screen "1121_OMACPackTags" 1280x715, template "1xxx_MachineControl"
   TextField "fraStatusPackTags" at 15,15 size 535x225; Text 'Status / Estado:'
   TextField "txtStatusCurUnitMode" at 25,55 size 220x25; Text 'Unit mode current: / Aktuelle Betriebsart: / Modo de unidad actual:'
   TextField "txtStatusCurState" at 25,85 size 220x25; Text 'State current: / Aktueller Zustand: / Corriente del estado'
   TextField "txtStatusCurMachSpeed" at 25,115 size 220x25; Text 'Current machine speed: / Aktuelle Geschwindigkeit'
   TextField "txtStatusCurMachSpeedUnit" at 370,115 size 80x25; Text 'pcs/min / Stck/Min / m/min'
   TextField "txtStatusMachSpeed" at 25,145 size 220x25; Text 'Machine speed: / Maschinengeschwindigkeit: / Velocidad de la máquina:'
   TextField "txtStatusMachSpeedUnit" at 370,145 size 80x25; Text 'pcs/min / Stck/Min / m/min'
   TextField "txtStatusEquipmentInterlockBlocked" at 25,175 size 220x25; Text 'Equip. interlock blocked: / Equip. interlock blockiert:'
   TextField "txtStatusEquipmentInterlockStarved" at 25,205 size 220x25; Text 'Equip. interlock starved: / Equip. interlock leer:'
   SymbolicIOField "valOutputStatusUnitMode" at 245,55 size 295x25; TextOn '1'; TextOff '0'; TextList "LPMLV30_UnitModes"
      ProcessValue <- "PackTags.Status.UnitModeCurrent"
   SymbolicIOField "valOutputStatusState" at 245,85 size 295x25; TextOn '1'; TextOff '0'; TextList "LPMLV30_States"
      ProcessValue <- "PackTags.Status.StateCurrent"
   IOField "valOutputStatusCurMachSpeed" at 245,115 size 125x25; FormatPattern 99999.9
      ProcessValue <- "PackTags.Status.CurMachSpeed"
   IOField "valOutputStatusMachSpeed" at 245,145 size 125x25; FormatPattern 99999.9
      ProcessValue <- "PackTags.Status.MachSpeed"
   IOField "valOutputStatusEquipmentInterlockBlocked" at 245,175 size 20x25; FormatPattern 1
      ProcessValue <- "PackTags.Status.EquipmentInterlock.Blocked"
   IOField "valOutputStatusEquipmentInterlockStarved" at 245,205 size 20x25; FormatPattern 1
      ProcessValue <- "PackTags.Status.EquipmentInterlock.Starved"
   TextField "fraCommandPackTags" at 555,15 size 535x225; Text 'Command'
   TextField "txtCommandMachSpeed" at 565,55 size 220x25; Text 'Machine speed: / Maschinengeschwindigkeit: / Velocidad de la máquina:'
   TextField "txtCommandMachSpeedUnit" at 910,55 size 80x25; Text 'pcs/min / Stck/Min / m/min'
   TextField "txtCommandUnitMode" at 565,85 size 220x25; Text 'Unit mode: / Modo de unidad:'
   TextField "txtCommandUnitModeChangeRequest" at 565,115 size 220x25; Text 'Mode change request:'
   TextField "txtCommandStateControl" at 565,145 size 220x25; Text 'State control command: / Comando de control del estado:'
   TextField "TxtCommandStateChangeRequest" at 565,175 size 220x25; Text 'State change request:'
   IOField "valOutputCommandMachSpeed" at 785,55 size 125x25; FormatPattern 99999.9
      ProcessValue <- "PackTags.Command.MachSpeed"
   SymbolicIOField "valOutputCommandUnitMode" at 785,85 size 295x25; TextOn '1'; TextOff '0'; TextList "LPMLV30_UnitModes"
      ProcessValue <- "PackTags.Command.UnitMode"
   IOField "valOutputCommandUnitModeChangeRequest" at 784,115 size 20x25; FormatPattern 1
      ProcessValue <- "PackTags.Command.UnitModeChangeRequest"
   SymbolicIOField "valOutputCommandStateControl" at 785,145 size 295x25; TextOn '1'; TextOff '0'; TextList "LPMLV30_States"
      ProcessValue <- "PackTags.Command.CntrlCmd"
   IOField "valOutputCommandStateControlChangeRequest" at 784,175 size 20x25; FormatPattern 1
      ProcessValue <- "PackTags.Command.CmdChangeRequest"
   TextField "fraAdminPackTags" at 15,245 size 1075x330; Text 'Admin'
   TextField "txtAdminCount" at 245,285 size 125x25; Text 'Counts / Zähler'
   TextField "txtAdminAccCount" at 375,285 size 125x25; Text 'Acc. Count / Akk. Zähler'
   TextField "txtAdminMachDesignSpeed" at 25,410 size 220x25; Text 'Machine design speed: / Sollgeschwindigkeit: / Velocidad de diseño de la máquina:'
   TextField "txtAdminMachDesignSpeedUnit" at 370,410 size 80x25; Text 'pcs/min / Stck/Min / m/min'
   TextField "txtAdminStopReasonID" at 25,450 size 220x25; Text 'Stop reason ID: / Detener identificación de la razón:'
   TextField "txtAdminStopReasonMessage" at 25,480 size 220x25; Text 'Stop reason message: / Fehlerursache: / Detener mensaje de motivo:'
   TextField "txtAdminActiveAlamrs" at 25,510 size 220x25; Text 'Active alarms: / Aktive Alarme:'
   TextField "txtAdminActiveWarnings" at 25,540 size 220x25; Text 'Active warnings: / Aktive Warnungen:'
   IOField "valOutputAdminConsumedCountName" at 25,310 size 220x25; FormatPattern ????????????????
      ProcessValue <- "PackTags.Admin.ProdConsumedCount[0].Name"
   IOField "valOutputAdminConsumedCountValue" at 245,310 size 125x25; FormatPattern s9999999999
      ProcessValue <- "PackTags.Admin.ProdConsumedCount[0].Count"
   IOField "valOutputAdminConsumedAccCountValue" at 375,310 size 125x25; FormatPattern s9999999999
      ProcessValue <- "PackTags.Admin.ProdConsumedCount[0].AccCount"
   IOField "valOutputAdminConsumedCountUnit" at 500,310 size 80x25; FormatPattern ??????
      ProcessValue <- "PackTags.Admin.ProdConsumedCount[0].Unit"
   IOField "valOutputAdminProcessedCountName" at 25,340 size 220x25; FormatPattern ????????????????
      ProcessValue <- "PackTags.Admin.ProdProcessedCount[0].Name"
   IOField "valOutputAdminProcessedCountValue" at 245,340 size 125x25; FormatPattern s9999999999
      ProcessValue <- "PackTags.Admin.ProdProcessedCount[0].Count"
   IOField "valOutputAdminProcessedAccCountValue" at 375,340 size 125x25; FormatPattern s9999999999
      ProcessValue <- "PackTags.Admin.ProdProcessedCount[0].AccCount"
   IOField "valOutputAdminProcessedCountUnit" at 500,340 size 80x25; FormatPattern ??????
      ProcessValue <- "PackTags.Admin.ProdProcessedCount[0].Unit"
   IOField "valOutputAdminDefectiveCountName" at 25,370 size 220x25; FormatPattern ????????????????
      ProcessValue <- "PackTags.Admin.ProdDefectiveCount[0].Name"
   IOField "valOutputAdminDefectiveCountValue" at 245,370 size 125x25; FormatPattern s9999999999
      ProcessValue <- "PackTags.Admin.ProdDefectiveCount[0].Count"
   IOField "valOutputAdminDefectiveAccCountValue" at 375,370 size 125x25; FormatPattern s9999999999
      ProcessValue <- "PackTags.Admin.ProdDefectiveCount[0].AccCount"
   IOField "valOutputAdminDefectiveCountUnit" at 500,370 size 80x25; FormatPattern ??????
      ProcessValue <- "PackTags.Admin.ProdDefectiveCount[0].Unit"
   IOField "valOutputAdminMachDesignSpeed" at 245,410 size 125x25; FormatPattern 9999.9
      ProcessValue <- "PackTags.Admin.MachDesignSpeed"
   IOField "valOutputAdminStopReasonID" at 245,450 size 125x25; FormatPattern 9999
      ProcessValue <- "PackTags.Admin.StopReason.ID"
   IOField "valOutputAdminStopReasonMessage" at 245,480 size 550x25; FormatPattern ????????????????????????????????????????????????????????????
      ProcessValue <- "PackTags.Admin.StopReason.Message"
   IOField "valOutputActiveAlarms" at 245,510 size 125x25; FormatPattern 99999
      ProcessValue <- "PackTags.Admin.AlarmExtent"
   IOField "valOutputActiveWarnings" at 245,540 size 125x25; FormatPattern 99999
      ProcessValue <- "PackTags.Admin.WarningExtent"
   Rectangle "recBaseScreenLocked" at 0,0 size 1280x708
      Visibility <- "bo_System_BaseScreenLocked"

screen "1161_OMACTimes" 1280x715, template "1xxx_MachineControl"
   TextField "fraModeTimes" at 15,15 size 535x200; Text 'Mode Times / Mode-Zeiten'
   TextField "txtModeName" at 50,80 size 150x25; Text 'Mode / Modo'
   TextField "txtModeLastTime" at 200,55 size 101x50; Text 'Last time [min] Letzte Zeit [min] Ultima vez'
   TextField "txtModeTotalTime" at 300,55 size 101x50; Text 'Total time [min] Gesamtzeit [min] Tiempo Total'
   TextField "txtModeTimeInMode" at 400,55 size 140x50; Text 'Time in mode [%] Zeit in Mode [%] % Tiempo en modo'
   Circle "valOutputMode1Active" at 27,109 size 18x18
      Visibility <- "PackTags.Status.UnitModeCurrent"
   Circle "valOutputMode2Active" at 27,134 size 18x18
      Visibility <- "PackTags.Status.UnitModeCurrent"
   Circle "valOutputMode3Active" at 27,159 size 18x18
      Visibility <- "PackTags.Status.UnitModeCurrent"
   Circle "valOutputMode4Active" at 27,184 size 18x18
      Visibility <- "PackTags.Status.UnitModeCurrent"
   ScreenModuleView "fcpTimesMode1" at 50,105 size 490x26; ScreenModuleType ""
      Guid_{11997190-50578} <- "[1]"
      Guid_{11997190-50584} <- "PackTags.Admin.ModeCumulativeTime[1]"
      Guid_{11997190-50582} <- "PackTags.Admin.ModeCurrentTime[1]"
      Guid_{11997190-50586} <- "PackTags.Admin.AccTimeSinceLastReset"
   ScreenModuleView "fcpTimesMode2" at 50,130 size 490x26; ScreenModuleType ""
      Guid_{11997190-50578} <- "[2]"
      Guid_{11997190-50584} <- "PackTags.Admin.ModeCumulativeTime[2]"
      Guid_{11997190-50582} <- "PackTags.Admin.ModeCurrentTime[2]"
      Guid_{11997190-50586} <- "PackTags.Admin.AccTimeSinceLastReset"
   ScreenModuleView "fcpTimesMode3" at 50,155 size 490x26; ScreenModuleType ""
      Guid_{11997190-50578} <- "[3]"
      Guid_{11997190-50584} <- "PackTags.Admin.ModeCumulativeTime[3]"
      Guid_{11997190-50582} <- "PackTags.Admin.ModeCurrentTime[3]"
      Guid_{11997190-50586} <- "PackTags.Admin.AccTimeSinceLastReset"
   ScreenModuleView "fcpTimesMode4" at 50,180 size 490x26; ScreenModuleType ""
      Guid_{11997190-50578} <- "[4]"
      Guid_{11997190-50584} <- "PackTags.Admin.ModeCumulativeTime[4]"
      Guid_{11997190-50582} <- "PackTags.Admin.ModeCurrentTime[4]"
      Guid_{11997190-50586} <- "PackTags.Admin.AccTimeSinceLastReset"
   TextField "txtTimeSinceLastReset" at 25,510 size 220x25; Text 'Time since last reset: / Zeit seit letztem Reset: / Tiempo desde el último reinicio:'
   TextField "txtTimeSinceLastResetUnit" at 369,510 size 80x25; Text 'min / min.'
   IOField "valOutputTimeSinceLastReset" at 244,510 size 125x25; FormatPattern 9999999999
      ProcessValue <- "PackTags.Admin.AccTimeSinceLastReset"
   Button "btnResetTimes" at 420,510 size 125x25; TextOff 'Reset / Restablecer temporizadores'
      on Release: ResetBit("HMI_Data.resetPackMLTimers")
      on Press: SetBit("HMI_Data.resetPackMLTimers")
      Appearance <- "HMI_Data.resetPackMLTimers"
   TextField "fraStateTimesOfCurrentMode" at 555,15 size 535x525; Text 'State Times of current Mode / State-Zeiten in aktuellem Mode'
   TextField "txtStateName" at 590,80 size 150x25; Text 'State / Modo'
   TextField "txtStateLastTime" at 740,55 size 101x50; Text 'Last time [min] Letzte Zeit [min] Ultima vez'
   TextField "txtStateTotalTime" at 840,55 size 101x50; Text 'Total time [min] Gesamtzeit [min] Tiempo Total'
   TextField "txtStateTimeInState" at 940,55 size 140x50; Text 'Time in state [%] Zeit in State [%] % Tiempo en modo'
   Circle "valOutputState1Active" at 567,109 size 18x18
      Visibility <- "PackTags.Status.StateCurrent"
   Circle "valOutputState2Active" at 567,134 size 18x18
      Visibility <- "PackTags.Status.StateCurrent"
   Circle "valOutputState3Active" at 567,159 size 18x18
      Visibility <- "PackTags.Status.StateCurrent"
   Circle "valOutputState4Active" at 567,184 size 18x18
      Visibility <- "PackTags.Status.StateCurrent"
   Circle "valOutputState5Active" at 567,209 size 18x18
      Visibility <- "PackTags.Status.StateCurrent"
   Circle "valOutputState6Active" at 567,234 size 18x18
      Visibility <- "PackTags.Status.StateCurrent"
   Circle "valOutputState7Active" at 567,259 size 18x18
      Visibility <- "PackTags.Status.StateCurrent"
   Circle "valOutputState8Active" at 567,284 size 18x18
      Visibility <- "PackTags.Status.StateCurrent"
   Circle "valOutputState9Active" at 567,309 size 18x18
      Visibility <- "PackTags.Status.StateCurrent"
   Circle "valOutputState10Active" at 567,335 size 18x18
      Visibility <- "PackTags.Status.StateCurrent"
   Circle "valOutputState11Active" at 567,359 size 18x18
      Visibility <- "PackTags.Status.StateCurrent"
   Circle "valOutputState12Active" at 567,384 size 18x18
      Visibility <- "PackTags.Status.StateCurrent"
   Circle "valOutputState13Active" at 567,409 size 18x18
      Visibility <- "PackTags.Status.StateCurrent"
   Circle "valOutputState14Active" at 567,434 size 18x18
      Visibility <- "PackTags.Status.StateCurrent"
   Circle "valOutputState15Active" at 567,459 size 18x18
      Visibility <- "PackTags.Status.StateCurrent"
   Circle "valOutputState16Active" at 567,484 size 18x18
      Visibility <- "PackTags.Status.StateCurrent"
   Circle "valOutputState17Active" at 567,509 size 18x18
      Visibility <- "PackTags.Status.StateCurrent"
   ScreenModuleView "fcpTimesState1" at 590,105 size 490x26; ScreenModuleType ""
      Guid_{11997190-50578} <- "[1]"
      Guid_{11997190-50584} <- "HMI_Data.State_Cumulative_Times[1]"
      Guid_{11997190-50582} <- "HMI_Data.State_Current_Times[1]"
      Guid_{11997190-50586} <- "HMI_Data.modeCumulativeTime"
   ScreenModuleView "fcpTimesState2" at 590,130 size 490x26; ScreenModuleType ""
      Guid_{11997190-50578} <- "[2]"
      Guid_{11997190-50584} <- "HMI_Data.State_Cumulative_Times[2]"
      Guid_{11997190-50582} <- "HMI_Data.State_Current_Times[2]"
      Guid_{11997190-50586} <- "HMI_Data.modeCumulativeTime"
   ScreenModuleView "fcpTimesState3" at 590,155 size 490x26; ScreenModuleType ""
      Guid_{11997190-50578} <- "[3]"
      Guid_{11997190-50584} <- "HMI_Data.State_Cumulative_Times[3]"
      Guid_{11997190-50582} <- "HMI_Data.State_Current_Times[3]"
      Guid_{11997190-50586} <- "HMI_Data.modeCumulativeTime"
   ScreenModuleView "fcpTimesState4" at 590,180 size 490x26; ScreenModuleType ""
      Guid_{11997190-50578} <- "[4]"
      Guid_{11997190-50584} <- "HMI_Data.State_Cumulative_Times[4]"
      Guid_{11997190-50582} <- "HMI_Data.State_Current_Times[4]"
      Guid_{11997190-50586} <- "HMI_Data.modeCumulativeTime"
   ScreenModuleView "fcpTimesState5" at 590,205 size 490x26; ScreenModuleType ""
      Guid_{11997190-50578} <- "[5]"
      Guid_{11997190-50584} <- "HMI_Data.State_Cumulative_Times[5]"
      Guid_{11997190-50582} <- "HMI_Data.State_Current_Times[5]"
      Guid_{11997190-50586} <- "HMI_Data.modeCumulativeTime"
   ScreenModuleView "fcpTimesState6" at 590,230 size 490x26; ScreenModuleType ""
      Guid_{11997190-50578} <- "[6]"
      Guid_{11997190-50584} <- "HMI_Data.State_Cumulative_Times[6]"
      Guid_{11997190-50582} <- "HMI_Data.State_Current_Times[6]"
      Guid_{11997190-50586} <- "HMI_Data.modeCumulativeTime"
   ScreenModuleView "fcpTimesState7" at 590,255 size 490x26; ScreenModuleType ""
      Guid_{11997190-50578} <- "[7]"
      Guid_{11997190-50584} <- "HMI_Data.State_Cumulative_Times[7]"
      Guid_{11997190-50582} <- "HMI_Data.State_Current_Times[7]"
      Guid_{11997190-50586} <- "HMI_Data.modeCumulativeTime"
   ScreenModuleView "fcpTimesState8" at 590,280 size 490x26; ScreenModuleType ""
      Guid_{11997190-50578} <- "[8]"
      Guid_{11997190-50584} <- "HMI_Data.State_Cumulative_Times[8]"
      Guid_{11997190-50582} <- "HMI_Data.State_Current_Times[8]"
      Guid_{11997190-50586} <- "HMI_Data.modeCumulativeTime"
   ScreenModuleView "fcpTimesState9" at 590,305 size 490x26; ScreenModuleType ""
      Guid_{11997190-50578} <- "[9]"
      Guid_{11997190-50584} <- "HMI_Data.State_Cumulative_Times[9]"
      Guid_{11997190-50582} <- "HMI_Data.State_Current_Times[9]"
      Guid_{11997190-50586} <- "HMI_Data.modeCumulativeTime"
   ScreenModuleView "fcpTimesState10" at 590,330 size 490x26; ScreenModuleType ""
      Guid_{11997190-50578} <- "[10]"
      Guid_{11997190-50584} <- "HMI_Data.State_Cumulative_Times[10]"
      Guid_{11997190-50582} <- "HMI_Data.State_Current_Times[10]"
      Guid_{11997190-50586} <- "HMI_Data.modeCumulativeTime"
   ScreenModuleView "fcpTimesState11" at 590,355 size 490x26; ScreenModuleType ""
      Guid_{11997190-50578} <- "[11]"
      Guid_{11997190-50584} <- "HMI_Data.State_Cumulative_Times[11]"
      Guid_{11997190-50582} <- "HMI_Data.State_Current_Times[11]"
      Guid_{11997190-50586} <- "HMI_Data.modeCumulativeTime"
   ScreenModuleView "fcpTimesState12" at 590,380 size 490x26; ScreenModuleType ""
      Guid_{11997190-50578} <- "[12]"
      Guid_{11997190-50584} <- "HMI_Data.State_Cumulative_Times[12]"
      Guid_{11997190-50582} <- "HMI_Data.State_Current_Times[12]"
      Guid_{11997190-50586} <- "HMI_Data.modeCumulativeTime"
   ScreenModuleView "fcpTimesState13" at 590,405 size 490x26; ScreenModuleType ""
      Guid_{11997190-50578} <- "[13]"
      Guid_{11997190-50584} <- "HMI_Data.State_Cumulative_Times[13]"
      Guid_{11997190-50582} <- "HMI_Data.State_Current_Times[13]"
      Guid_{11997190-50586} <- "HMI_Data.modeCumulativeTime"
   ScreenModuleView "fcpTimesState14" at 590,430 size 490x26; ScreenModuleType ""
      Guid_{11997190-50578} <- "[14]"
      Guid_{11997190-50584} <- "HMI_Data.State_Cumulative_Times[14]"
      Guid_{11997190-50582} <- "HMI_Data.State_Current_Times[14]"
      Guid_{11997190-50586} <- "HMI_Data.modeCumulativeTime"
   ScreenModuleView "fcpTimesState15" at 590,455 size 490x26; ScreenModuleType ""
      Guid_{11997190-50578} <- "[15]"
      Guid_{11997190-50584} <- "HMI_Data.State_Cumulative_Times[15]"
      Guid_{11997190-50582} <- "HMI_Data.State_Current_Times[15]"
      Guid_{11997190-50586} <- "HMI_Data.modeCumulativeTime"
   ScreenModuleView "fcpTimesState16" at 590,480 size 490x26; ScreenModuleType ""
      Guid_{11997190-50578} <- "[16]"
      Guid_{11997190-50584} <- "HMI_Data.State_Cumulative_Times[16]"
      Guid_{11997190-50582} <- "HMI_Data.State_Current_Times[16]"
      Guid_{11997190-50586} <- "HMI_Data.modeCumulativeTime"
   ScreenModuleView "fcpTimesState17" at 590,505 size 490x26; ScreenModuleType ""
      Guid_{11997190-50578} <- "[17]"
      Guid_{11997190-50584} <- "HMI_Data.State_Cumulative_Times[17]"
      Guid_{11997190-50582} <- "HMI_Data.State_Current_Times[17]"
      Guid_{11997190-50586} <- "HMI_Data.modeCumulativeTime"
   Rectangle "recBaseScreenLocked" at 0,0 size 1280x708
      Visibility <- "bo_System_BaseScreenLocked"

screen "1241_ManualCommands" 1280x715, template "1xxx_MachineControl"
   Button "btnEnableRemoteChangeCmd" at 90,175 size 125x275; TextOff 'Reset / Reiniciar'; TextList "Local_Remote_Control"; PictureOff "Start_gray_32x32"
      on Release: InvertBit("PackML.remoteCommandEnable")
      Appearance <- "PackML.remoteCommandEnable"
      ProcessValue <- "PackML.remoteCommandEnable"
   Rectangle "valOutputLocalChangeCmdEnabled" at 220,175 size 795x165
      Visibility <- "PackML.remoteCommandEnable"
   TextField "fraLocalChangeCmd" at 220,175 size 795x165; Text 'Local Change Commands / Comandos de control de modo / Lokale Kommandos'
   Button "btnLocalChangeCmdProduction" at 230,225 size 125x50; TextOff 'Production / Produktion / Produccion'
      on Release: ResetBit("PackML.Cmd.Mode.Production")
      on Press: SetBit("PackML.Cmd.Mode.Production")
      Appearance <- "PackML.Cmd.Mode.Production"
      ObjectEnable <- "PackML.remoteCommandEnable"
   Button "btnLocalChangeCmdMaintenance" at 360,225 size 125x50; TextOff 'Maintenance / Wartung / Manual'
      on Release: ResetBit("PackML.Cmd.Mode.Maintenance")
      on Press: SetBit("PackML.Cmd.Mode.Maintenance")
      Appearance <- "PackML.Cmd.Mode.Maintenance"
      ObjectEnable <- "PackML.remoteCommandEnable"
   Button "btnLocalChangeCmdManual" at 490,225 size 125x50; TextOff 'Manual / Jog / Hand / Tippen / Manual'
      on Release: ResetBit("PackML.Cmd.Mode.Manual")
      on Press: SetBit("PackML.Cmd.Mode.Manual")
      Appearance <- "PackML.Cmd.Mode.Manual"
      ObjectEnable <- "PackML.remoteCommandEnable"
   Button "btnLocalChangeCmdUserMode1" at 620,225 size 125x50; TextOff 'User Mode 1 Benutzer- mode 1 Manual'
      on Release: ResetBit("PackML.Cmd.Mode.UserMode01")
      on Press: SetBit("PackML.Cmd.Mode.UserMode01")
      Appearance <- "PackML.Cmd.Mode.UserMode01"
      ObjectEnable <- "PackML.remoteCommandEnable"
   Button "btnLocalChangeCmdStart" at 230,280 size 125x50; TextOff 'Start / Comienzo'
      on Release: ResetBit("HMI_Data.CMDs.PB_Start")
      on Press: SetBit("HMI_Data.CMDs.PB_Start")
      Appearance <- "HMI_Data.CMDs.PB_Start"
      ObjectEnable <- "PackML.remoteCommandEnable"
   Button "btnLocalChangeCmdStop" at 360,280 size 125x50; TextOff 'Stop / Detener'
      on Release: ResetBit("HMI_Data.CMDs.PB_Stop")
      on Press: SetBit("HMI_Data.CMDs.PB_Stop")
      Appearance <- "HMI_Data.CMDs.PB_Stop"
      ObjectEnable <- "PackML.remoteCommandEnable"
   Button "btnLocalChangeCmdReset" at 490,280 size 125x50; TextOff 'Reset / Reiniciar'
      on Release: ResetBit("HMI_Data.CMDs.PB_Reset")
      on Press: SetBit("HMI_Data.CMDs.PB_Reset")
      Appearance <- "HMI_Data.CMDs.PB_Reset"
      ObjectEnable <- "PackML.remoteCommandEnable"
   Button "btnLocalChangeCmdHold" at 620,280 size 125x50; TextOff 'Hold'
      on Release: ResetBit("HMI_Data.CMDs.PB_Hold")
      on Press: SetBit("HMI_Data.CMDs.PB_Hold")
      Appearance <- "HMI_Data.CMDs.PB_Hold"
      ObjectEnable <- "PackML.remoteCommandEnable"
   Button "btnLocalChangeCmdAbort" at 750,280 size 125x50; TextOff 'Abort'
      on Release: ResetBit("HMI_Data.CMDs.PB_Abort")
      on Press: SetBit("HMI_Data.CMDs.PB_Abort")
      Appearance <- "HMI_Data.CMDs.PB_Abort"
      ObjectEnable <- "PackML.remoteCommandEnable"
   Button "btnLocalChangeCmdComplete" at 880,280 size 125x50; TextOff 'Complete'
      on Release: ResetBit("HMI_Data.CMDs.PB_Complete")
      on Press: SetBit("HMI_Data.CMDs.PB_Complete")
      Appearance <- "HMI_Data.CMDs.PB_Complete"
      ObjectEnable <- "PackML.remoteCommandEnable"
   Rectangle "valOutputRemoteChangeCmdEnabled" at 220,345 size 795x105
      Visibility <- "PackML.remoteCommandEnable"
   TextField "fraRemoteChangeCmd" at 220,345 size 795x105; Text 'Remote Change Commands / Comando de control del estado: / Remote Kommandos'
   TextField "txtRemoteModeChangeCmd" at 355,385 size 220x25; Text 'Mode change command: / Mode-Wechsel: / Comando de cambio de modo remoto:'
   TextField "txtRemoteStateChangeCmd" at 356,415 size 220x25; Text 'State change command: / State-Wechsel: / Comando de cambio de modo remoto:'
   SymbolicIOField "valInputRemoteModeChangeCmd" at 575,385 size 300x25; TextOn '1'; TextOff '0'; TextList "LPMLV30_UnitModes"
      Appearance <- "PackML.remoteCommandEnable"
      ProcessValue <- "PackTags.Command.UnitMode"
      ObjectEnable <- "PackML.remoteCommandEnable"
   SymbolicIOField "valInputRemoteStateChangeCmd" at 575,415 size 300x25; TextOn '1'; TextOff '0'; TextList "LPMLV30_CntrlCmd"
      Appearance <- "PackML.remoteCommandEnable"
      ProcessValue <- "PackTags.Command.CntrlCmd"
      ObjectEnable <- "PackML.remoteCommandEnable"
   Button "btnRemoteModeChangeCmdConfirm" at 880,385 size 125x25; TextOn 'Text Comando de control Habilitado'; TextOff 'Confirm Übernehmen Comando de control Discapacitado'; PictureOff "Start_gray_32x32"
      on Release: ResetBit("PackTags.Command.UnitModeChangeRequest")
      on Press: SetBit("PackTags.Command.UnitModeChangeRequest")
      Appearance <- "PackTags.Command.UnitModeChangeRequest"
      ObjectEnable <- "PackML.remoteCommandEnable"
   Button "btnRemoteStateChangeCmdConfirm" at 880,415 size 125x25; TextOn 'Text Comando de control Habilitado'; TextOff 'Confirm Übernehmen Comando de control Discapacitado'; PictureOff "Start_gray_32x32"
      on Release: ResetBit("PackTags.Command.CmdChangeRequest")
      on Press: SetBit("PackTags.Command.CmdChangeRequest")
      Appearance <- "PackTags.Command.CmdChangeRequest"
      ObjectEnable <- "PackML.remoteCommandEnable"
   Rectangle "recBaseScreenLocked" at 0,0 size 1280x708
      Visibility <- "bo_System_BaseScreenLocked"

screen "1201_OEE" 1280x715, template "1xxx_MachineControl"
   TextField "fraModeTimes" at 15,15 size 1075x277; Text 'Overall Equipment Effectiveness / Gesamtanlageneffektivität'
   Gauge "valOutputGaugeOEE" at 70,70 size 220x220; CaptionText 'Overall OEE / Gesamt OEE'; UnitText 'Unit'
      ProcessValue <- "PackML.OEE.realTime"
   Gauge "valOutputGaugeAvailablity" at 310,70 size 220x220; CaptionText 'Availability / Verfügbarkeit'; UnitText 'Unit'
      ProcessValue <- "PackML.OEE.availability"
   Gauge "valOutputGaugePerformance" at 550,70 size 220x220; CaptionText 'Performance / Actuación / Leistung'; UnitText 'Unit'
      ProcessValue <- "PackML.OEE.performance"
   Gauge "valOutputGaugeQuality" at 790,70 size 220x220; CaptionText 'Quality / Qualität'; UnitText 'Unit'
      ProcessValue <- "PackML.OEE.quality"
   IOField "valOutputOEE" at 129,210 size 65x25; FormatPattern 999.9
      ProcessValue <- "PackML.OEE.realTime"
   IOField "valOutputAvailability" at 369,210 size 65x25; FormatPattern 999.9
      ProcessValue <- "PackML.OEE.availability"
   IOField "valOutputPerformance" at 609,210 size 65x25; FormatPattern 999.9
      ProcessValue <- "PackML.OEE.performance"
   IOField "valOutputQuality" at 849,210 size 65x25; FormatPattern 999.9
      ProcessValue <- "PackML.OEE.quality"
   TextField "txtOEEUnit" at 194,210 size 80x25; Text '%'
   TextField "txtAvailabiltyUnit" at 434,210 size 80x25; Text '%'
   TextField "txtPerformanceUnit" at 674,210 size 80x25; Text '%'
   TextField "txtQualityUnit" at 914,210 size 80x25; Text '%'
   Rectangle "recBaseScreenLocked" at 0,0 size 1280x708
      Visibility <- "bo_System_BaseScreenLocked"

screen "2041_SystemFunctions" 1280x715, template "2xxx_Settings"
   on GenerateScreen: function_ed885d1a("i16_Settings_CurDisplayBrightness")
   TextField "fraSystemTime" at 15,15 size 1075x80; Text 'System time / Systemzeit / hora del sistema'
   TextField "txtCurSystemTime" at 25,55 size 220x25; Text 'Current system time: / Aktuelle Systemzeit:'
   DateTimeField "valOutputCurSystemTime" at 245,55 size 230x25
   TextField "txtNewSystemTime" at 495,55 size 220x25; Text 'New system time: / Neue Systemzeit: / Nuevo tiempo del sistema:'
   DateTimeField "valInputNewSystemTime" at 715,55 size 230x25
      ProcessValue <- "dat_Settings_NewDateTime"
   Button "btnSetNewSystemTime" at 950,55 size 125x25; TextOff 'Confirm / Übernehmen'
   TextField "fraScreenBrightness" at 15,100 size 1075x110; Text 'Screen Brightness / Bildschirmhelligkeit'
   Bar "valOutput1ScreenBrightness" at 85,145 size 935x50; MinimumValue 0; MaximumValue 100
      ProcessValue <- "i16_Settings_CurDisplayBrightness"
   IOField "valOutput2ScreenBrightness" at 85,145 size 935x50; FormatPattern 999; Unit  %
      ProcessValue <- "i16_Settings_CurDisplayBrightness"
   Button "btnScreenBrightnessPlus" at 1025,145 size 50x50; TextOff '+'
      on Release: "sub_SetScreenBrightness"(10)
   Button "btnScreenBrightnessMinus" at 30,145 size 50x50; TextOff '-'
      on Release: "sub_SetScreenBrightness"(-10)
   TextField "txtLanguage" at 15,215 size 535x100; Text 'Language / Sprache / Idioma'
   Button "btnSelectEnglish" at 25,255 size 125x50; TextOff 'Text'; PictureOff "pic-flag-USA-201x134"
      on Click: function_fb9197e8(L en-US); SetTag("HMI_Data.languageSelected", 0)
   Button "btnSelectGerman" at 155,255 size 125x50; TextOff 'Text'; PictureOff "pic-flag-GE-201x134"
      on Click: function_fb9197e8(L de-DE); SetTag("HMI_Data.languageSelected", 1)
   TextField "txtSystemFunctions" at 555,215 size 535x100; Text 'Functions / Funktionen'
   Button "btnOpenScreenCleaning" at 565,255 size 125x50; TextOff 'Clean Screen Bildschirm- reinigung'
      on Release: function_be740847(30)
   Button "btnOpenTouchCalibrate" at 695,255 size 125x50; TextOff 'Touch Calibration Touch Kalibrierung Toque Calibración'
      on Release: function_bc3e350c()
   Button "btnRuntimeStop" at 825,255 size 125x50; TextOff 'Stop Runtime Runtime beenden Detener el tiempo de ejecución'
      on Release: StopRuntime(0)
   Rectangle "recBaseScreenLocked" at 0,0 size 1280x708
      Visibility <- "bo_System_BaseScreenLocked"
   Button "btnSelectSpain" at 285,255 size 125x50; TextOff 'Text'; PictureOff "SPAN001"
      on Click: function_fb9197e8(L en-US); SetTag("HMI_Data.languageSelected", 2)

screen "2081_UserManagement" 1280x715, template "2xxx_Settings"
   UserView "ctrlUserManagement" at 15,15 size 1035x480
      ObjectEnable <- "bo_System_BaseScreenLocked"
   Button "btnUserManagementVerticalScrollUp" at 1050,40 size 40x30; TextOff 'Text'; PictureOff "icn-scroll-up-20x11"
      on Release: function_b22acb07("ctrlUserManagement")
   Button "btnUserManagementVerticalScrollDown" at 1050,465 size 40x30; TextOff 'Text'; PictureOff "icn-scroll-down-20x11"
      on Release: function_b8b2ebe3("ctrlUserManagement")
   TextField "txtUserAccessInfo" at 15,500 size 272x109; Text 'User Access: 1) admin / admin (full access) 2) simatic / simatic (full access) 3) maint / maint (limited access) 4) user / user (basic access) User Acces: 1) admin / admin (full access) 2) simatic / simatic (full access) 3) maint / maint (limited access) 4) user / user (basic access)'
   Rectangle "recBaseScreenLocked" at 0,0 size 1280x708
      Visibility <- "bo_System_BaseScreenLocked"

screen "2001_Settings" 1280x715, template "2xxx_Settings"
   Button "rec_BaseScreenLocked" at 0,0 size 1280x715; TextOff 'Text'
      Visibility <- "bo_System_BaseScreenLocked"

screen "3001_AlarmOverview" 1280x715, template "3xxx_Alarms&Events"
   TextField "fraStopReasonAlarmHistory" at 15,245 size 1075x175; Text 'Stop Reason Alarm History / Stop Reason Alarmhistory / Detener el historial de alarmas de la razón:'
   TextField "txtStopReasonAlarmHistoryID" at 50,285 size 55x25; Text 'ID / ID:'
   TextField "txtStopReasonAlarmHistoryValue" at 105,285 size 55x25; Text 'Value / Valor:'
   TextField "txtStopReasonAlarmHistoryCategory" at 160,285 size 30x25; Text 'Cat / Kat'
   TextField "txtStopReasonAlarmHistoryMessage" at 190,285 size 490x25; Text 'Message / Meldung / Mensaje:'
   TextField "txtStopReasonAlarmHistoryTimeIn" at 680,285 size 200x25; Text 'Time In / Gekommen / Tiempo en:'
   TextField "txtStopReasonAlarmHistoryTimeOut" at 880,285 size 200x25; Text 'Time Out / Gegangen / Se acabó el tiempo:'
   TextField "txtStopReasonAlarmHistoryRow1" at 25,310 size 25x25; Text '1'
   TextField "txtStopReasonAlarmHistoryRow2" at 25,335 size 25x25; Text '2'
   TextField "txtStopReasonAlarmHistoryRow3" at 25,360 size 25x25; Text '3'
   TextField "txtStopReasonAlarmHistoryRow4" at 25,385 size 25x25; Text '4'
   ScreenModuleView "fcpStopReasonAlarmHistoryRow1-2" at 50,310 size 1030x51; ScreenModuleType ""
      Guid_{11997190-460713} <- "PackTags.Admin.AlarmHistory[1]"
      Guid_{11997190-460693} <- "PackTags.Admin.AlarmHistory[0]"
   ScreenModuleView "fcpStopReasonAlarmHistoryRow3-4" at 50,360 size 1030x51; ScreenModuleType ""
      Guid_{11997190-460713} <- "PackTags.Admin.AlarmHistory[3]"
      Guid_{11997190-460693} <- "PackTags.Admin.AlarmHistory[2]"
   TextField "fraActiveWarnings" at 15,425 size 1075x175; Text 'Active Warnings / Aktive Warnungen'
   TextField "txtActiveWarningsID" at 50,465 size 55x25; Text 'ID / ID:'
   TextField "txtActiveWarningsCategory" at 105,465 size 30x25; Text 'Cat / Kat'
   TextField "txtActiveWarningsMessage" at 135,465 size 545x25; Text 'Message / Meldung / Mensaje:'
   TextField "txtActiveWarningsTimeIn" at 680,465 size 200x25; Text 'Time In / Gekommen / Tiempo en:'
   TextField "txtActiveWarningsTimeOut" at 880,465 size 200x25; Text 'Time Out / Gegangen / Se acabó el tiempo:'
   TextField "txtActiveWarningsRow1" at 25,490 size 25x25; Text '1'
   TextField "txtActiveWarningsRow2" at 25,515 size 25x25; Text '2'
   TextField "txtActiveWarningsRow3" at 25,540 size 25x25; Text '3'
   TextField "txtActiveWarningsRow4" at 25,565 size 25x25; Text '4'
   ScreenModuleView "fcpActiveWarningsRow1-2" at 50,490 size 1030x51; ScreenModuleType ""
      Guid_{11997190-460713} <- "HMI_Data.warningSortedList[1]"
      Guid_{11997190-460693} <- "HMI_Data.warningSortedList[0]"
   ScreenModuleView "fcpActiveWarningsRow3-4" at 50,540 size 1030x51; ScreenModuleType ""
      Guid_{11997190-460713} <- "HMI_Data.warningSortedList[3]"
      Guid_{11997190-460693} <- "HMI_Data.warningSortedList[2]"
   TextField "fraActiveAlarms" at 15,15 size 1075x225; Text 'Active Alarms / Aktive Alarme'
   TextField "txtActiveAlarmsID" at 50,55 size 55x25; Text 'ID / ID:'
   TextField "txtActiveAlarmsValue" at 105,55 size 55x25; Text 'Value / Valor:'
   TextField "txtActiveAlarmsCategory" at 160,55 size 30x25; Text 'Cat / Kat'
   TextField "txtActiveAlarmsMessage" at 190,55 size 490x25; Text 'Message / Meldung / Mensaje:'
   TextField "txtActiveAlarmsTimeIn" at 680,55 size 200x25; Text 'Time In / Gekommen / Tiempo en:'
   TextField "txtActiveAlarmsTimeOut" at 880,55 size 200x25; Text 'Time Out / Gegangen / Se acabó el tiempo:'
   TextField "txtActiveAlarmsRow1" at 25,80 size 25x25; Text '1'
   TextField "txtActiveAlarmsRow2" at 25,105 size 25x25; Text '2'
   TextField "txtActiveAlarmsRow3" at 25,130 size 25x25; Text '3'
   TextField "txtActiveAlarmsRow4" at 25,155 size 25x25; Text '4'
   TextField "txtActiveAlarmsRow5" at 25,180 size 25x25; Text '5'
   TextField "txtActiveAlarmsRow6" at 25,205 size 25x25; Text '6'
   ScreenModuleView "fcpActiveAlarmsRow1-2" at 50,80 size 1030x51; ScreenModuleType ""
      Guid_{11997190-460713} <- "HMI_Data.alarmSortedList[1]"
      Guid_{11997190-460693} <- "HMI_Data.alarmSortedList[0]"
   ScreenModuleView "fcpActiveAlarmsRow3-4" at 50,130 size 1030x51; ScreenModuleType ""
      Guid_{11997190-460713} <- "HMI_Data.alarmSortedList[3]"
      Guid_{11997190-460693} <- "HMI_Data.alarmSortedList[2]"
   ScreenModuleView "fcpActiveAlarmsRow5-6" at 50,180 size 1030x51; ScreenModuleType ""
      Guid_{11997190-460713} <- "HMI_Data.alarmSortedList[5]"
      Guid_{11997190-460693} <- "HMI_Data.alarmSortedList[4]"
   Rectangle "recBaseScreenLocked" at 0,0 size 1280x708
      Visibility <- "bo_System_BaseScreenLocked"

screen "3041_AlarmEvents" 1280x715, template "3xxx_Alarms&Events"
   TextField "txtFilterCategory" at 180,55 size 250x25; Text 'Category: / Kategorie:'
   SymbolicIOField "valInputFilterCategory" at 180,80 size 250x25; TextOn '1'; TextOff '0'; TextList "CPG_CategoryList"
      Appearance <- "HMI_Data.alarmFilter.cmdFilterCategory"
      ProcessValue <- "HMI_Data.alarmFilter.cfgFilterCategory"
      ObjectEnable <- "HMI_Data.alarmFilter.cmdFilterCategory"
   Button "btnFilterCatagory" at 50,55 size 125x50; TextOff 'Filter Category Filter Kategorie Filtrar Categoría'
      on Release: InvertBit("HMI_Data.alarmFilter.cmdFilterCategory")
      Appearance <- "HMI_Data.alarmFilter.cmdFilterCategory"
   Button "btnFilterActiveEvents" at 435,55 size 125x50; TextOff 'Filter Active Events Filter aktive Meldungen Filtro activo Eventos'
      on Release: InvertBit("HMI_Data.alarmFilter.cmdFilterActiveEvents")
      Appearance <- "HMI_Data.alarmFilter.cmdFilterActiveEvents"
   Button "btnFilterUnit" at 15,560 size 125x50; TextOff 'Unit'
      on Release: InvertBit("HMI_Data.EM_SortDisable_Alarm.Unit")
      Appearance <- "HMI_Data.EM_SortDisable_Alarm.Unit"
      Visibility <- "UN.PackML_Sts.moduleActive"
   Button "btnFilterEM00" at 145,560 size 125x50; TextOff 'EM00 General Fct EM00 Zentrale Fkt EM00 Virtual EM'
      on Release: InvertBit("HMI_Data.EM_SortDisable_Alarm.EM00")
      Visibility <- "EM00.PackML_Sts.Unit.moduleActive"
      Appearance <- "HMI_Data.EM_SortDisable_Alarm.EM00"
   Button "btnFilterEM01" at 275,560 size 125x50; TextOff 'EM01'
      on Release: InvertBit("HMI_Data.EM_SortDisable_Alarm.EM01")
      Visibility <- "EM01.PackML_Sts.Unit.moduleActive"
      Appearance <- "HMI_Data.EM_SortDisable_Alarm.EM01"
   Button "btnFilterEM02" at 405,560 size 125x50; TextOff 'EM02'
      on Release: InvertBit("HMI_Data.EM_SortDisable_Alarm.EM02")
      Appearance <- "HMI_Data.EM_SortDisable_Alarm.EM02"
      Visibility <- "EM02.PackML_Sts.Unit.moduleActive"
   Button "btnSortByCategory" at 825,55 size 125x50; TextOff 'Sort by Category Sortieren nach Kategorie Sort by Category'
      on Release: InvertBit("HMI_Data.alarmFilter.cfgTimeSortDirection")
      Appearance <- "HMI_Data.alarmFilter.cfgTimeSortDirection"
   Button "btnSortByTime" at 955,55 size 125x50; TextOff 'Sort by Time Sortieren nach Zeit Ordenar por Hora'
      on Release: InvertBit("HMI_Data.alarmFilter.cmdSortCategory")
      Appearance <- "HMI_Data.alarmFilter.cmdSortCategory"
   TextField "fraAlarmEvents" at 15,15 size 1075x535; Text 'Alarm Events / Alarmmeldungen'
   TextField "txtAlarmEventsID" at 50,115 size 55x25; Text 'ID / ID:'
   TextField "txtAlarmEventsValue" at 105,115 size 55x25; Text 'Value / Valor:'
   TextField "txtAlarmEventsCategory" at 160,115 size 30x25; Text 'Cat / Kat'
   TextField "txtAlarmEventsMessage" at 190,115 size 490x25; Text 'Message / Meldung / Mensaje:'
   TextField "txtAlarmEventsTimeIn" at 680,115 size 200x25; Text 'Time In / Gekommen / Tiempo en:'
   TextField "txtAlarmEventsTimeOut" at 880,115 size 200x25; Text 'Time Out / Gegangen / Se acabó el tiempo:'
   TextField "txtAlarmEventsRow1" at 25,140 size 25x25; Text '1'
   TextField "txtAlarmEventsRow2" at 25,165 size 25x25; Text '2'
   TextField "txtAlarmEventsRow3" at 25,190 size 25x25; Text '3'
   TextField "txtAlarmEventsRow4" at 25,215 size 25x25; Text '4'
   TextField "txtAlarmEventsRow5" at 25,240 size 25x25; Text '5'
   TextField "txtAlarmEventsRow6" at 25,265 size 25x25; Text '6'
   TextField "txtAlarmEventsRow7" at 25,290 size 25x25; Text '7'
   TextField "txtAlarmEventsRow8" at 25,315 size 25x25; Text '8'
   TextField "txtAlarmEventsRow9" at 25,340 size 25x25; Text '9'
   TextField "txtAlarmEventsRow10" at 25,365 size 25x25; Text '10'
   TextField "txtAlarmEventsRow11" at 25,390 size 25x25; Text '11'
   TextField "txtAlarmEventsRow12" at 25,415 size 25x25; Text '12'
   TextField "txtAlarmEventsRow13" at 25,440 size 25x25; Text '13'
   TextField "txtAlarmEventsRow14" at 25,465 size 25x25; Text '14'
   TextField "txtAlarmEventsRow15" at 25,490 size 25x25; Text '15'
   TextField "txtAlarmEventsRow16" at 25,515 size 25x25; Text '16'
   ScreenModuleView "fcpAlarmEventsRow1-2" at 50,140 size 1030x51; ScreenModuleType ""
      Guid_{11997190-460713} <- "HMI_Data.alarmSortedList[1]"
      Guid_{11997190-460693} <- "HMI_Data.alarmSortedList[0]"
   ScreenModuleView "fcpAlarmEventsRow3-4" at 50,190 size 1030x51; ScreenModuleType ""
      Guid_{11997190-460713} <- "HMI_Data.alarmSortedList[3]"
      Guid_{11997190-460693} <- "HMI_Data.alarmSortedList[2]"
   ScreenModuleView "fcpAlarmEventsRow5-6" at 50,240 size 1030x51; ScreenModuleType ""
      Guid_{11997190-460713} <- "HMI_Data.alarmSortedList[5]"
      Guid_{11997190-460693} <- "HMI_Data.alarmSortedList[4]"
   ScreenModuleView "fcpAlarmEventsRow7-8" at 50,290 size 1030x51; ScreenModuleType ""
      Guid_{11997190-460713} <- "HMI_Data.alarmSortedList[7]"
      Guid_{11997190-460693} <- "HMI_Data.alarmSortedList[6]"
   ScreenModuleView "fcpAlarmEventsRow9-10" at 50,340 size 1030x51; ScreenModuleType ""
      Guid_{11997190-460713} <- "HMI_Data.alarmSortedList[9]"
      Guid_{11997190-460693} <- "HMI_Data.alarmSortedList[8]"
   ScreenModuleView "fcpAlarmEventsRow11-12" at 50,390 size 1030x51; ScreenModuleType ""
      Guid_{11997190-460713} <- "HMI_Data.alarmSortedList[11]"
      Guid_{11997190-460693} <- "HMI_Data.alarmSortedList[10]"
   ScreenModuleView "fcpAlarmEventsRow13-14" at 50,440 size 1030x51; ScreenModuleType ""
      Guid_{11997190-460713} <- "HMI_Data.alarmSortedList[13]"
      Guid_{11997190-460693} <- "HMI_Data.alarmSortedList[12]"
   ScreenModuleView "fcpAlarmEventsRow15-16" at 50,490 size 1030x51; ScreenModuleType ""
      Guid_{11997190-460713} <- "HMI_Data.alarmSortedList[15]"
      Guid_{11997190-460693} <- "HMI_Data.alarmSortedList[14]"
   Rectangle "recBaseScreenLocked" at 0,0 size 1280x708
      Visibility <- "bo_System_BaseScreenLocked"

screen "3081_WarningEvents" 1280x715, template "3xxx_Alarms&Events"
   TextField "txtFilterCategory" at 180,55 size 250x25; Text 'Category: / Kategorie:'
   SymbolicIOField "valInputFilterCategory" at 180,80 size 250x25; TextOn '1'; TextOff '0'; TextList "CPG_CategoryList"
      Appearance <- "HMI_Data.alarmFilter.cmdFilterCategory"
      ObjectEnable <- "HMI_Data.alarmFilter.cmdFilterCategory"
      ProcessValue <- "HMI_Data.alarmFilter.cfgFilterCategory"
   Button "btnFilterCatagory" at 50,55 size 125x50; TextOff 'Filter Category Filter Kategorie Filtrar Categoría'
      on Release: InvertBit("HMI_Data.alarmFilter.cmdFilterCategory")
      Appearance <- "HMI_Data.alarmFilter.cmdFilterCategory"
   Button "btnFilterActiveEvents" at 435,55 size 125x50; TextOff 'Filter Active Events Filter aktive Meldungen Filtro activo Eventos'
      on Release: InvertBit("HMI_Data.alarmFilter.cmdFilterActiveEvents")
      Appearance <- "HMI_Data.alarmFilter.cmdFilterActiveEvents"
   Button "btnFilterUnit" at 15,560 size 125x50; TextOff 'Unit'
      on Release: InvertBit("HMI_Data.EMSortDisableWarning.Unit")
      Appearance <- "HMI_Data.EMSortDisableWarning.Unit"
      Visibility <- "UN.PackML_Sts.moduleActive"
   Button "btnFilterEM00" at 145,560 size 125x50; TextOff 'EM00 General Fct EM00 Zentrale Fkt EM00 Virtual EM'
      on Release: InvertBit("HMI_Data.EMSortDisableWarning.EM00")
      Visibility <- "EM00.PackML_Sts.Unit.moduleActive"
      Appearance <- "HMI_Data.EMSortDisableWarning.EM00"
   Button "btnFilterEM01" at 275,560 size 125x50; TextOff 'EM01'
      on Release: InvertBit("HMI_Data.EMSortDisableWarning.EM01")
      Visibility <- "EM01.PackML_Sts.Unit.moduleActive"
      Appearance <- "HMI_Data.EMSortDisableWarning.EM01"
   Button "btnFilterEM02" at 405,560 size 125x50; TextOff 'EM02'
      on Release: InvertBit("HMI_Data.EMSortDisableWarning.EM02")
      Appearance <- "HMI_Data.EMSortDisableWarning.EM02"
      Visibility <- "EM02.PackML_Sts.Unit.moduleActive"
   Button "btnSortByCategory" at 825,55 size 125x50; TextOff 'Sort by Category Sortieren nach Kategorie Ordenar por Categoría'
      on Release: InvertBit("HMI_Data.alarmFilter.cfgTimeSortDirection")
      Appearance <- "HMI_Data.alarmFilter.cfgTimeSortDirection"
   Button "btnSortByTime" at 955,55 size 125x50; TextOff 'Sort by Time Sortieren nach Zeit Ordenar por Hora'
      on Release: InvertBit("HMI_Data.alarmFilter.cmdSortCategory")
      Appearance <- "HMI_Data.alarmFilter.cmdSortCategory"
   TextField "fraWarningEvents" at 15,15 size 1075x535; Text 'Warning Events / Warnungen'
   TextField "txtWarningEventsID" at 50,115 size 55x25; Text 'ID / ID:'
   TextField "txtWarningEventsCategory" at 105,115 size 30x25; Text 'Cat / Kat'
   TextField "txtWarningEventsMessage" at 135,115 size 545x25; Text 'Message / Meldung / Mensaje:'
   TextField "txtWarningEventsTimeIn" at 680,115 size 200x25; Text 'Time In / Gekommen / Tiempo en:'
   TextField "txtWarningEventsTimeOut" at 880,115 size 200x25; Text 'Time Out / Gegangen / Se acabó el tiempo:'
   TextField "txtWarningEventsRow1" at 25,140 size 25x25; Text '1'
   TextField "txtWarningEventsRow2" at 25,165 size 25x25; Text '2'
   TextField "txtWarningEventsRow3" at 25,190 size 25x25; Text '3'
   TextField "txtWarningEventsRow4" at 25,215 size 25x25; Text '4'
   TextField "txtWarningEventsRow5" at 25,240 size 25x25; Text '5'
   TextField "txtWarningEventsRow6" at 25,265 size 25x25; Text '6'
   TextField "txtWarningEventsRow7" at 25,290 size 25x25; Text '7'
   TextField "txtWarningEventsRow8" at 25,315 size 25x25; Text '8'
   TextField "txtWarningEventsRow9" at 25,340 size 25x25; Text '9'
   TextField "txtWarningEventsRow10" at 25,365 size 25x25; Text '10'
   TextField "txtWarningEventsRow11" at 25,390 size 25x25; Text '11'
   TextField "txtWarningEventsRow12" at 25,415 size 25x25; Text '12'
   TextField "txtWarningEventsRow13" at 25,440 size 25x25; Text '13'
   TextField "txtWarningEventsRow14" at 25,465 size 25x25; Text '14'
   TextField "txtWarningEventsRow15" at 25,490 size 25x25; Text '15'
   TextField "txtWarningEventsRow16" at 25,515 size 25x25; Text '16'
   ScreenModuleView "fcpWarningEventsRow1-2" at 50,190 size 1030x51; ScreenModuleType ""
      Guid_{11997190-460713} <- "HMI_Data.warningSortedList[3]"
      Guid_{11997190-460693} <- "HMI_Data.warningSortedList[2]"
   ScreenModuleView "fcpWarningEventsRow3-4" at 50,140 size 1030x51; ScreenModuleType ""
      Guid_{11997190-460713} <- "HMI_Data.warningSortedList[1]"
      Guid_{11997190-460693} <- "HMI_Data.warningSortedList[0]"
   ScreenModuleView "fcpWarningEventsRow5-6" at 50,240 size 1030x51; ScreenModuleType ""
      Guid_{11997190-460713} <- "HMI_Data.warningSortedList[5]"
      Guid_{11997190-460693} <- "HMI_Data.warningSortedList[4]"
   ScreenModuleView "fcpWarningEventsRow7-8" at 50,290 size 1030x51; ScreenModuleType ""
      Guid_{11997190-460713} <- "HMI_Data.warningSortedList[7]"
      Guid_{11997190-460693} <- "HMI_Data.warningSortedList[6]"
   ScreenModuleView "fcpWarningEventsRow9-10" at 50,340 size 1030x51; ScreenModuleType ""
      Guid_{11997190-460713} <- "HMI_Data.warningSortedList[9]"
      Guid_{11997190-460693} <- "HMI_Data.warningSortedList[8]"
   ScreenModuleView "fcpWarningEventsRow11-12" at 50,390 size 1030x51; ScreenModuleType ""
      Guid_{11997190-460713} <- "HMI_Data.warningSortedList[11]"
      Guid_{11997190-460693} <- "HMI_Data.warningSortedList[10]"
   ScreenModuleView "fcpWarningEventsRow13-14" at 50,440 size 1030x51; ScreenModuleType ""
      Guid_{11997190-460713} <- "HMI_Data.warningSortedList[13]"
      Guid_{11997190-460693} <- "HMI_Data.warningSortedList[12]"
   ScreenModuleView "fcpWarningEventsRow15-16" at 50,490 size 1030x51; ScreenModuleType ""
      Guid_{11997190-460713} <- "HMI_Data.warningSortedList[15]"
      Guid_{11997190-460693} <- "HMI_Data.warningSortedList[14]"
   Rectangle "recBaseScreenLocked" at 0,0 size 1280x708
      Visibility <- "bo_System_BaseScreenLocked"

screen "3121_HMI_Alarms" 1280x715, template "3xxx_Alarms&Events"
   TextField "fraHMIMessageHistory" at 15,315 size 1075x295; Text 'HMI Events History / HMI Meldehistorie / Alarmas y advertencias borradas'
   AlarmView "ctrlHMIMessageHistory" at 25,355 size 1015x245; ColumnTextAlarmText 'Text / Texto'; AlarmLog "Message Archive"
      ObjectEnable <- "bo_System_BaseScreenLocked"
   Button "btnHMIMessageHistoryVerticalScrollUp" at 1040,381 size 40x30; TextOff 'Text'; PictureOff "icn-scroll-up-20x11"
      on Release: function_b22acb07("ctrlHMIMessageHistory")
   Button "btnHMIMessageHistoryVerticalScrollDown" at 1040,570 size 40x30; TextOff 'Text'; PictureOff "icn-scroll-down-20x11"
      on Release: function_b8b2ebe3("ctrlHMIMessageHistory")
   TextField "fraActiveHMIMessages" at 15,15 size 1075x295; Text 'Active HMI Events / Aktive HMI Meldungen: / Alarmas activas y advertencias'
   AlarmView "ctrlActiveHMIMessages" at 25,55 size 1015x245; ColumnTextAlarmText 'Text / Texto'
      ObjectEnable <- "bo_System_BaseScreenLocked"
   Button "btnActiveHMIMessagesVerticalScrollUp" at 1040,81 size 40x30; TextOff 'Text'; PictureOff "icn-scroll-up-20x11"
      on Release: function_b22acb07("ctrlActiveHMIMessages")
   Button "btnActiveHMIMessagesVerticalScrollDown" at 1040,270 size 40x30; TextOff 'Text'; PictureOff "icn-scroll-down-20x11"
      on Release: function_b8b2ebe3("ctrlActiveHMIMessages")
   Rectangle "recBaseScreenLocked" at 0,0 size 1280x708
      Visibility <- "bo_System_BaseScreenLocked"